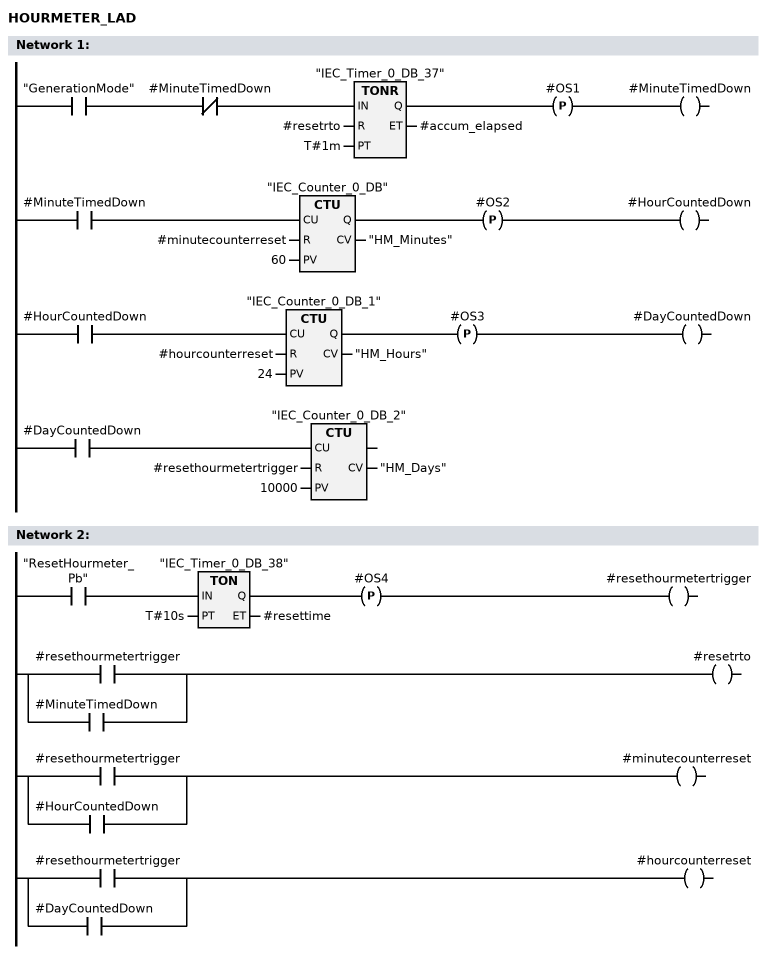
   "IEC_Timer_0_DB_37".TONR(IN := "GenerationMode" AND NOT #MinuteTimedDown,
                           R := #resetrto,
                           PT := T#1m,
                           ET => #accum_elapsed);
   #_w1 := "IEC_Timer_0_DB_37".Q AND NOT #OS1;   // rising edge
   #OS1 := "IEC_Timer_0_DB_37".Q;
   #MinuteTimedDown := #_w1;
   "IEC_Counter_0_DB".CTU(CU := #MinuteTimedDown, R := #minutecounterreset, PV := 60, CV => "HM_Minutes");
   #_w2 := "IEC_Counter_0_DB".Q AND NOT #OS2;   // rising edge
   #OS2 := "IEC_Counter_0_DB".Q;
   #HourCountedDown := #_w2;
   "IEC_Counter_0_DB_1".CTU(CU := #HourCountedDown, R := #hourcounterreset, PV := 24, CV => "HM_Hours");
   #_w3 := "IEC_Counter_0_DB_1".Q AND NOT #OS3;   // rising edge
   #OS3 := "IEC_Counter_0_DB_1".Q;
   #DayCountedDown := #_w3;
   "IEC_Counter_0_DB_2".CTU(CU := #DayCountedDown, R := #resethourmetertrigger, PV := 10000, CV => "HM_Days");
END_REGION

REGION Network 2
   "IEC_Timer_0_DB_38".TON(IN := "ResetHourmeter_Pb", PT := T#10s, ET => #resettime);
   #_w1 := "IEC_Timer_0_DB_38".Q AND NOT #OS4;   // rising edge
   #OS4 := "IEC_Timer_0_DB_38".Q;
   #resethourmetertrigger := #_w1;
   #resetrto := #resethourmetertrigger OR #MinuteTimedDown;
   #minutecounterreset := #resethourmetertrigger OR #HourCountedDown;
   #hourcounterreset := #resethourmetertrigger OR #DayCountedDown;
END_REGION
END_FUNCTION_BLOCK

FUNCTION_BLOCK "HOURMETER_FBD"   // FB20, FBD
{ S7_Optimized_Access := 'TRUE' }
VERSION : 0.1
   VAR
      OS1 : Bool;
      OS2 : Bool;
      OS3 : Bool;
      OS4 : Bool;
      rtotimerreset : Bool;
      minutecounterreset : Bool;
      hourcounterreset : Bool;
      hourmeterresettrigger : Bool;
      accumulatedtime : Time;
      minutetimeddown : Bool;
      hourcounteddown : Bool;
      daycounteddown : Bool;
   END_VAR
   VAR_TEMP   // added for the SCL form of the ladder/FBD networks
      _w1 : Bool;
      _w2 : Bool;
      _w3 : Bool;
   END_VAR
BEGIN

REGION Network 1
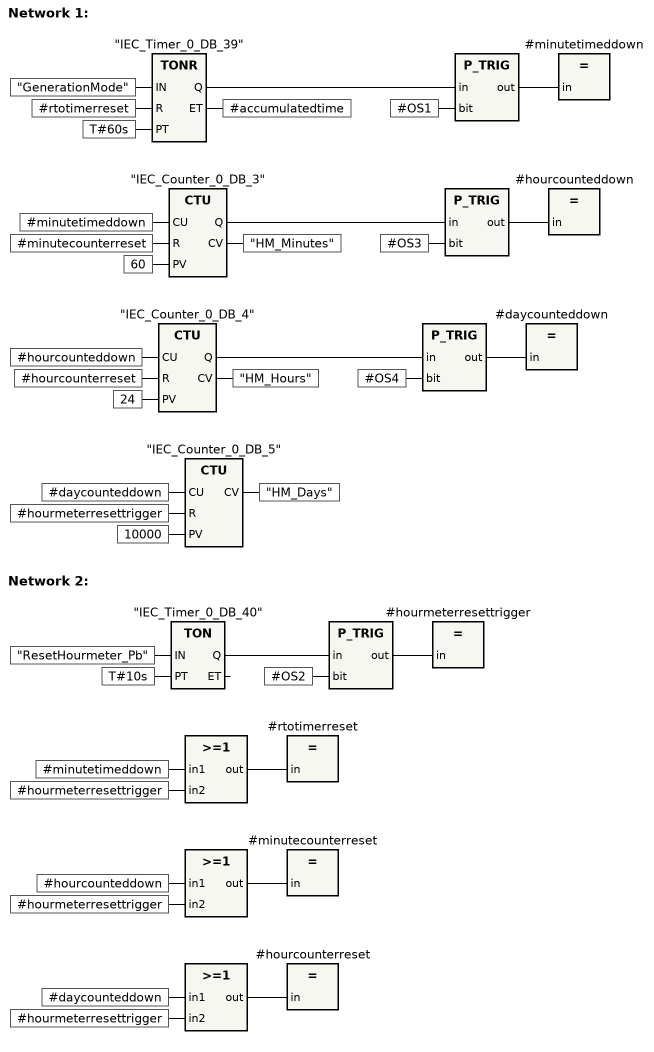
   "IEC_Timer_0_DB_39".TONR(IN := "GenerationMode", R := #rtotimerreset, PT := T#60s, ET => #accumulatedtime);
   #_w1 := "IEC_Timer_0_DB_39".Q AND NOT #OS1;   // rising edge
   #OS1 := "IEC_Timer_0_DB_39".Q;
   #minutetimeddown := #_w1;
   "IEC_Counter_0_DB_3".CTU(CU := #minutetimeddown, R := #minutecounterreset, PV := 60, CV => "HM_Minutes");
   #_w2 := "IEC_Counter_0_DB_3".Q AND NOT #OS3;   // rising edge
   #OS3 := "IEC_Counter_0_DB_3".Q;
   #hourcounteddown := #_w2;
   "IEC_Counter_0_DB_4".CTU(CU := #hourcounteddown, R := #hourcounterreset, PV := 24, CV => "HM_Hours");
   #_w3 := "IEC_Counter_0_DB_4".Q AND NOT #OS4;   // rising edge
   #OS4 := "IEC_Counter_0_DB_4".Q;
   #daycounteddown := #_w3;
   "IEC_Counter_0_DB_5".CTU(CU := #daycounteddown, R := #hourmeterresettrigger, PV := 10000, CV => "HM_Days");
END_REGION

REGION Network 2
   "IEC_Timer_0_DB_40".TON(IN := "ResetHourmeter_Pb", PT := T#10s);
   #_w1 := "IEC_Timer_0_DB_40".Q AND NOT #OS2;   // rising edge
   #OS2 := "IEC_Timer_0_DB_40".Q;
   #hourmeterresettrigger := #_w1;
   #rtotimerreset := #minutetimeddown OR #hourmeterresettrigger;
   #minutecounterreset := #hourcounteddown OR #hourmeterresettrigger;
   #hourcounterreset := #daycounteddown OR #hourmeterresettrigger;
END_REGION
END_FUNCTION_BLOCK

FUNCTION_BLOCK "HOURMETER_SCL"   // FB21, SCL
{ S7_Optimized_Access := 'TRUE' }
VERSION : 0.1
   VAR
      rtotimerreset : Bool;
      minutecounterreset : Bool;
      hourcounterreset : Bool;
      hourmeterresettrigger : Bool;
      accumulatedtime : Time;
      minutetimeddown : Bool;
      hourcounteddown : Bool;
      daycounteddown : Bool;
   END_VAR
BEGIN
   IF "GenerationMode" THEN
       "IEC_Timer_0_DB_41".TONR(IN := TRUE,
                                R := #rtotimerreset,
                                PT := T#60s,
                                Q => #minutetimeddown,
                                ET => #accumulatedtime);
   END_IF;

   IF #minutetimeddown THEN
       RESET_TIMER("IEC_Timer_0_DB_41");
   END_IF;

   "IEC_Counter_0_DB_6".CTU(CU:=#minutetimeddown,
                            R:=#minutecounterreset,
                            PV:=60,
                            Q=>#hourcounteddown,
                            CV=>"HM_Minutes");

   "IEC_Counter_0_DB_7".CTU(CU:=#hourcounteddown,
                            R:=#hourcounterreset,
                            PV:=24,
                            Q=>#daycounteddown,
                            CV=>"HM_Hours");

   "IEC_Counter_0_DB_9".CTU(CU:=#daycounteddown,
                            R:=#hourmeterresettrigger,
                            PV:=10000,
                            CV=>"HM_Days");

   IF "ResetHourmeter_Pb" THEN
       "IEC_Timer_0_DB_42".TON(IN:=TRUE,
                               PT:=T#10s,
                               Q=>#hourmeterresettrigger);
   ELSE
       RESET_TIMER("IEC_Timer_0_DB_42");
   END_IF;

   IF #hourmeterresettrigger OR #minutetimeddown THEN
       #rtotimerreset := 1;
   ELSE
       #rtotimerreset := 0;
   END_IF;

   IF #hourmeterresettrigger OR #hourcounteddown THEN
       #minutecounterreset := 1;
   ELSE
       #minutecounterreset := 0;
   END_IF;

   IF #hourmeterresettrigger OR #daycounteddown THEN
       #hourcounterreset := 1;
   ELSE
       #hourcounterreset := 0;
   END_IF;
END_FUNCTION_BLOCK

FUNCTION_BLOCK "HOURMETER_STL"   // FB22, STL
{ S7_Optimized_Access := 'TRUE' }
VERSION : 0.1
   VAR
      hourmeterresettrigger : Bool;
      minutecounterreset : Bool;
      hourcounterreset : Bool;
      minutetimeddown : Bool;
      hourcounteddown : Bool;
      daycounteddown : Bool;
      accumulatedtime : Time;
      rtotimerreset : Bool;
   END_VAR
   VAR_TEMP
      toomanydays : Bool;
      acctime : Time;
   END_VAR
BEGIN

REGION Network 1
         A     "GenerationMode";
         JC    RTOtimer;
         CLR;
         JU    EndOfLine;

   RTOtimer:CALL  TONR, "IEC_Timer_0_DB_43"
         ( IN := TRUE,
           R  := #rtotimerreset,
           PT := T#1m,
           Q  := #minutetimeddown,
           ET := #accumulatedtime
         );

         CALL  CTU, "IEC_Counter_0_DB_10"
         ( CU := #minutetimeddown,
           R  := #minutecounterreset,
           PV := 60,
           Q  := #hourcounteddown,
           CV := "HM_Minutes"
         );

         CALL  CTU, "IEC_Counter_0_DB_11"
         ( CU := #hourcounteddown,
           R  := #hourcounterreset,
           PV := 24,
           Q  := #daycounteddown,
           CV := "HM_Hours"
         );

         CALL  CTU, "IEC_Counter_0_DB_12"
         ( CU := #daycounteddown,
           R  := #hourmeterresettrigger,
           PV := 10000,
           Q  := #toomanydays,
           CV := "HM_Days"
         );

         JU    ResetEvaluate;

   ResetEvaluate:CLR;
         A     "ResetHourmeter_Pb";
         JC    ResetHourmeter;
         CALL  RESET_TIMER
         ( "TIMER" := "IEC_Timer_0_DB_44"
         );
         JU    EndOfLine;

   ResetHourmeter:CALL  TON, "IEC_Timer_0_DB_44"
         ( IN := TRUE,
           PT := T#10s,
           Q  := #hourmeterresettrigger,
           ET := #acctime
         );


   EndOfLine:A     #hourmeterresettrigger;
         O     #minutetimeddown;
         =     #rtotimerreset;
         CLR;
         A     #hourmeterresettrigger;
         O     #hourcounteddown;
         =     #minutecounterreset;
         CLR;
         A     #hourmeterresettrigger;
         O     #daycounteddown;
         =     #hourcounterreset;
         CLR;
         NOT;
         R     #hourmeterresettrigger;
END_REGION
END_FUNCTION_BLOCK

FUNCTION "SCP" : Void   // FC1, FBD
{ S7_Optimized_Access := 'TRUE' }
VERSION : 0.1
   VAR_INPUT
      Input_Min : Int;
      Input_Signal : Int;
      Input_Max : Int;
      Output_Min : Int;
      Output_Max : Int;
   END_VAR
   VAR_OUTPUT
      SV : Int;
   END_VAR
   VAR_TEMP
      tv : Real;
   END_VAR
BEGIN

REGION Network 1
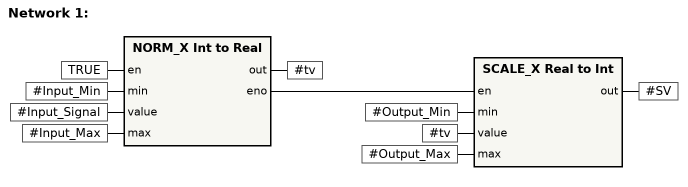
   IF TRUE THEN
       #tv := NORM_X(MIN := #Input_Min, VALUE := #Input_Signal, MAX := #Input_Max);
       #SV := SCALE_X(MIN := #Output_Min, VALUE := #tv, MAX := #Output_Max);
   END_IF;
END_REGION
END_FUNCTION

FUNCTION "CONVERTTIME" : Void   // FC2, FBD
{ S7_Optimized_Access := 'TRUE' }
VERSION : 0.1
   VAR_INPUT
      Int1 : Int;
   END_VAR
   VAR_OUTPUT
      Time1 : Time;
   END_VAR
   VAR_TEMP
      tv : Int;
   END_VAR
BEGIN

REGION Network 1
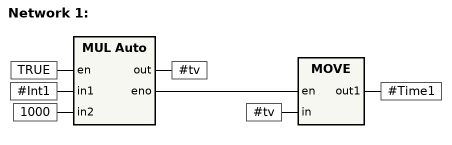
   IF TRUE THEN
       #tv := #Int1 * 1000;
       #Time1 := #tv;
   END_IF;
END_REGION
END_FUNCTION

ORGANIZATION_BLOCK "Main"   // OB1, LAD, ProgramCycle
TITLE = "Main Program Sweep (Cycle)"
{ S7_Optimized_Access := 'TRUE' }
VERSION : 0.1
   VAR_INPUT
      Initial_Call : Bool;   // Initial call of this OB
      Remanence : Bool;   // =True, if remanent data are available
   END_VAR
   VAR_TEMP
      SequenceInit : Bool;
      InitSequence : Bool;
   END_VAR
   VAR_TEMP   // added for the SCL form of the ladder/FBD networks
      _w1 : Bool;
      _w2 : Bool;
      _w3 : Bool;
      _w4 : Bool;
   END_VAR
BEGIN

REGION Network 1
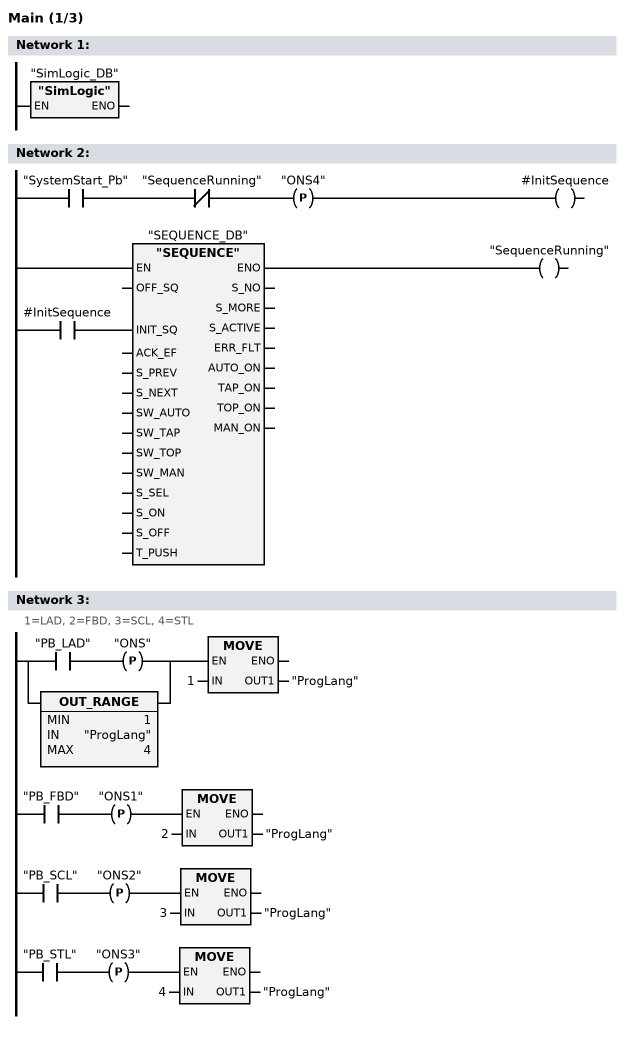
   RUNG wire#powerrail
      "SimLogic_DB"()
   END_RUNG
   // the same network as SCL:
   "SimLogic_DB"();   // "SimLogic"
END_REGION

REGION Network 2
   RUNG wire#powerrail
      Contact( "SystemStart_Pb" )
      I_Contact( "SequenceRunning" )
      P_Trig( "ONS4" )
      Coil( #InitSequence )
   END_RUNG
   RUNG wire#powerrail
      "SEQUENCE_DB"(INIT_SQ := wire#w1, OFF_SQ :=, ACK_EF :=, S_PREV :=, S_NEXT :=, SW_AUTO :=, SW_TAP :=, SW_TOP :=, SW_MAN :=, S_SEL :=, S_ON :=, S_OFF :=, T_PUSH :=, S_NO =>, S_MORE =>, S_ACTIVE =>, ERR_FLT =>, AUTO_ON =>, TAP_ON =>, TOP_ON =>, MAN_ON =>)
      Coil( "SequenceRunning" )
   END_RUNG
   RUNG wire#powerrail
      Contact( #InitSequence )
   END_RUNG wire#w1
   // the same network as SCL:
   #_w1 := "SystemStart_Pb" AND NOT "SequenceRunning";
   #_w2 := #_w1 AND NOT "ONS4";   // rising edge
   "ONS4" := #_w1;
   #InitSequence := #_w2;
   "SEQUENCE_DB"(INIT_SQ := #InitSequence, ENO => #_w3);   // "SEQUENCE"
   "SequenceRunning" := #_w3;
END_REGION

REGION Network 3
   // 1=LAD, 2=FBD, 3=SCL, 4=STL
   #_w1 := "PB_LAD" AND NOT "ONS";   // rising edge
   "ONS" := "PB_LAD";
   IF #_w1 OR ("ProgLang" < 1) OR ("ProgLang" > 4) THEN "ProgLang" := 1; END_IF;
   #_w2 := "PB_FBD" AND NOT "ONS1";   // rising edge
   "ONS1" := "PB_FBD";
   IF #_w2 THEN "ProgLang" := 2; END_IF;
   #_w3 := "PB_SCL" AND NOT "ONS2";   // rising edge
   "ONS2" := "PB_SCL";
   IF #_w3 THEN "ProgLang" := 3; END_IF;
   #_w4 := "PB_STL" AND NOT "ONS3";   // rising edge
   "ONS3" := "PB_STL";
   IF #_w4 THEN "ProgLang" := 4; END_IF;
END_REGION

REGION Network 4
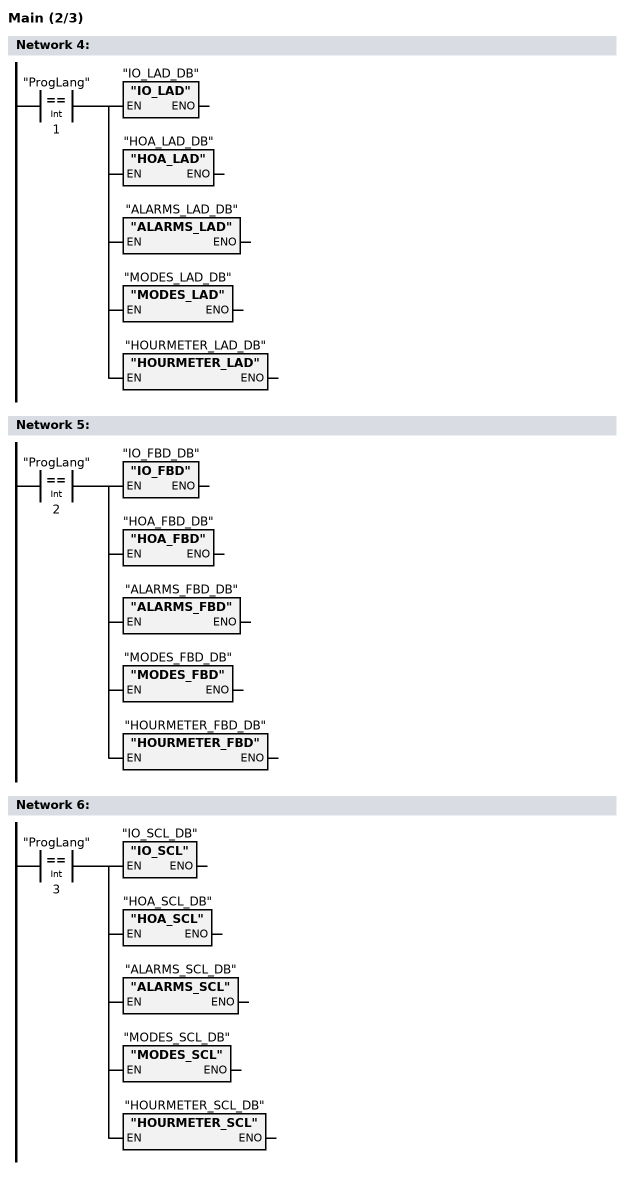
   RUNG wire#powerrail
      { S7_Templates := "SrcType := Int" } EQ_Contact(in1 := "ProgLang", in2 := 1)
      wire#w1
      "IO_LAD_DB"()
   END_RUNG
   RUNG wire#w1
      "HOA_LAD_DB"()
   END_RUNG
   RUNG wire#w1
      "ALARMS_LAD_DB"()
   END_RUNG
   RUNG wire#w1
      "MODES_LAD_DB"()
   END_RUNG
   RUNG wire#w1
      "HOURMETER_LAD_DB"()
   END_RUNG
   // the same network as SCL:
   #_w1 := "ProgLang" = 1;
   IF #_w1 THEN
       "IO_LAD_DB"();   // "IO_LAD"
       "HOA_LAD_DB"();   // "HOA_LAD"
       "ALARMS_LAD_DB"();   // "ALARMS_LAD"
       "MODES_LAD_DB"();   // "MODES_LAD"
       "HOURMETER_LAD_DB"();   // "HOURMETER_LAD"
   END_IF;
END_REGION

REGION Network 5
   RUNG wire#powerrail
      { S7_Templates := "SrcType := Int" } EQ_Contact(in1 := "ProgLang", in2 := 2)
      wire#w1
      "IO_FBD_DB"()
   END_RUNG
   RUNG wire#w1
      "HOA_FBD_DB"()
   END_RUNG
   RUNG wire#w1
      "ALARMS_FBD_DB"()
   END_RUNG
   RUNG wire#w1
      "MODES_FBD_DB"()
   END_RUNG
   RUNG wire#w1
      "HOURMETER_FBD_DB"()
   END_RUNG
   // the same network as SCL:
   #_w1 := "ProgLang" = 2;
   IF #_w1 THEN
       "IO_FBD_DB"();   // "IO_FBD"
       "HOA_FBD_DB"();   // "HOA_FBD"
       "ALARMS_FBD_DB"();   // "ALARMS_FBD"
       "MODES_FBD_DB"();   // "MODES_FBD"
       "HOURMETER_FBD_DB"();   // "HOURMETER_FBD"
   END_IF;
END_REGION

REGION Network 6
   RUNG wire#powerrail
      { S7_Templates := "SrcType := Int" } EQ_Contact(in1 := "ProgLang", in2 := 3)
      wire#w1
      "IO_SCL_DB"()
   END_RUNG
   RUNG wire#w1
      "HOA_SCL_DB"()
   END_RUNG
   RUNG wire#w1
      "ALARMS_SCL_DB"()
   END_RUNG
   RUNG wire#w1
      "MODES_SCL_DB"()
   END_RUNG
   RUNG wire#w1
      "HOURMETER_SCL_DB"()
   END_RUNG
   // the same network as SCL:
   #_w1 := "ProgLang" = 3;
   IF #_w1 THEN
       "IO_SCL_DB"();   // "IO_SCL"
       "HOA_SCL_DB"();   // "HOA_SCL"
       "ALARMS_SCL_DB"();   // "ALARMS_SCL"
       "MODES_SCL_DB"();   // "MODES_SCL"
       "HOURMETER_SCL_DB"();   // "HOURMETER_SCL"
   END_IF;
END_REGION

REGION Network 7
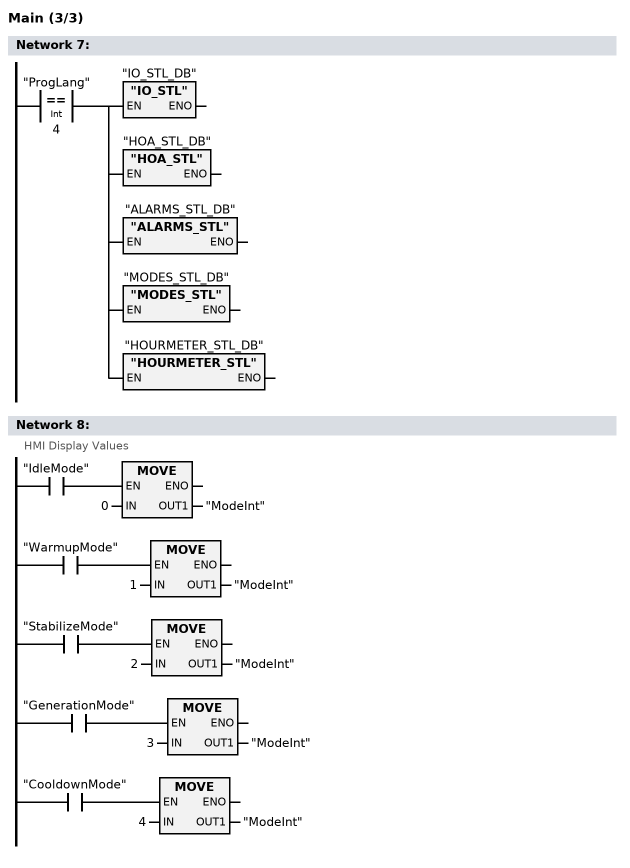
   RUNG wire#powerrail
      { S7_Templates := "SrcType := Int" } EQ_Contact(in1 := "ProgLang", in2 := 4)
      wire#w1
      "IO_STL_DB"()
   END_RUNG
   RUNG wire#w1
      "HOA_STL_DB"()
   END_RUNG
   RUNG wire#w1
      "ALARMS_STL_DB"()
   END_RUNG
   RUNG wire#w1
      "MODES_STL_DB"()
   END_RUNG
   RUNG wire#w1
      "HOURMETER_STL_DB"()
   END_RUNG
   // the same network as SCL:
   #_w1 := "ProgLang" = 4;
   IF #_w1 THEN
       "IO_STL_DB"();   // "IO_STL"
       "HOA_STL_DB"();   // "HOA_STL"
       "ALARMS_STL_DB"();   // "ALARMS_STL"
       "MODES_STL_DB"();   // "MODES_STL"
       "HOURMETER_STL_DB"();   // "HOURMETER_STL"
   END_IF;
END_REGION

REGION Network 8
   // HMI Display Values
   RUNG wire#powerrail
      Contact( "IdleMode" )
      Move(in := 0, out1 => "ModeInt")
   END_RUNG
   RUNG wire#powerrail
      Contact( "WarmupMode" )
      Move(in := 1, out1 => "ModeInt")
   END_RUNG
   RUNG wire#powerrail
      Contact( "StabilizeMode" )
      Move(in := 2, out1 => "ModeInt")
   END_RUNG
   RUNG wire#powerrail
      Contact( "GenerationMode" )
      Move(in := 3, out1 => "ModeInt")
   END_RUNG
   RUNG wire#powerrail
      Contact( "CooldownMode" )
      Move(in := 4, out1 => "ModeInt")
   END_RUNG
   // the same network as SCL:
   IF "IdleMode" THEN "ModeInt" := 0; END_IF;
   IF "WarmupMode" THEN "ModeInt" := 1; END_IF;
   IF "StabilizeMode" THEN "ModeInt" := 2; END_IF;
   IF "GenerationMode" THEN "ModeInt" := 3; END_IF;
   IF "CooldownMode" THEN "ModeInt" := 4; END_IF;
END_REGION
END_ORGANIZATION_BLOCK

ORGANIZATION_BLOCK "PID"   // OB31, LAD, CyclicInterrupt
{ S7_Optimized_Access := 'TRUE' }
VERSION : 0.1
   VAR_INPUT
      Initial_Call : Bool;   // Initial call of this OB
      Event_Count : Int;   // Events discarded
   END_VAR
   VAR_TEMP
      Bsp : Real;
      Vsp : Real;
      BaffleHandTrigger : Bool;
      BaffleOffTrigger : Bool;
      VFDHandTrigger : Bool;
      VFDOffTrigger : Bool;
      BaffleAutoTrigger : Bool;
      VFDautoTrigger : Bool;
   END_VAR
   VAR_TEMP   // added for the SCL form of the ladder/FBD networks
      _w1 : Bool;
      _w2 : Bool;
      _w3 : Bool;
      _w4 : Bool;
      _w5 : Bool;
      _w6 : Bool;
      _w7 : Bool;
   END_VAR
BEGIN

REGION Network 1
   // High Oil Flow Alarm Handling
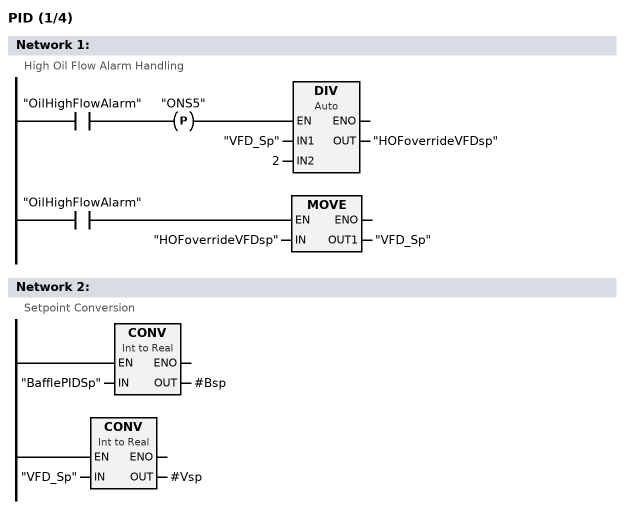
   RUNG wire#powerrail
      Contact( "OilHighFlowAlarm" )
      P_Trig( "ONS5" )
      Div(in1 := "VFD_Sp", in2 := 2, out => "HOFoverrideVFDsp")
   END_RUNG
   RUNG wire#powerrail
      Contact( "OilHighFlowAlarm" )
      Move(in := "HOFoverrideVFDsp", out1 => "VFD_Sp")
   END_RUNG
   // the same network as SCL:
   #_w1 := "OilHighFlowAlarm" AND NOT "ONS5";   // rising edge
   "ONS5" := "OilHighFlowAlarm";
   IF #_w1 THEN "HOFoverrideVFDsp" := "VFD_Sp" / 2; END_IF;
   IF "OilHighFlowAlarm" THEN "VFD_Sp" := "HOFoverrideVFDsp"; END_IF;
END_REGION

REGION Network 2
   // Setpoint Conversion
   RUNG wire#powerrail
      { S7_Templates := "[SrcType := Int, DestType := Real]" } Convert(in := "BafflePIDSp", out => #Bsp)
   END_RUNG
   RUNG wire#powerrail
      { S7_Templates := "[SrcType := Int, DestType := Real]" } Convert(in := "VFD_Sp", out => #Vsp)
   END_RUNG
   // the same network as SCL:
   #Bsp := INT_TO_REAL("BafflePIDSp");
   #Vsp := INT_TO_REAL("VFD_Sp");
END_REGION

REGION Network 3
   // Baffle HOA
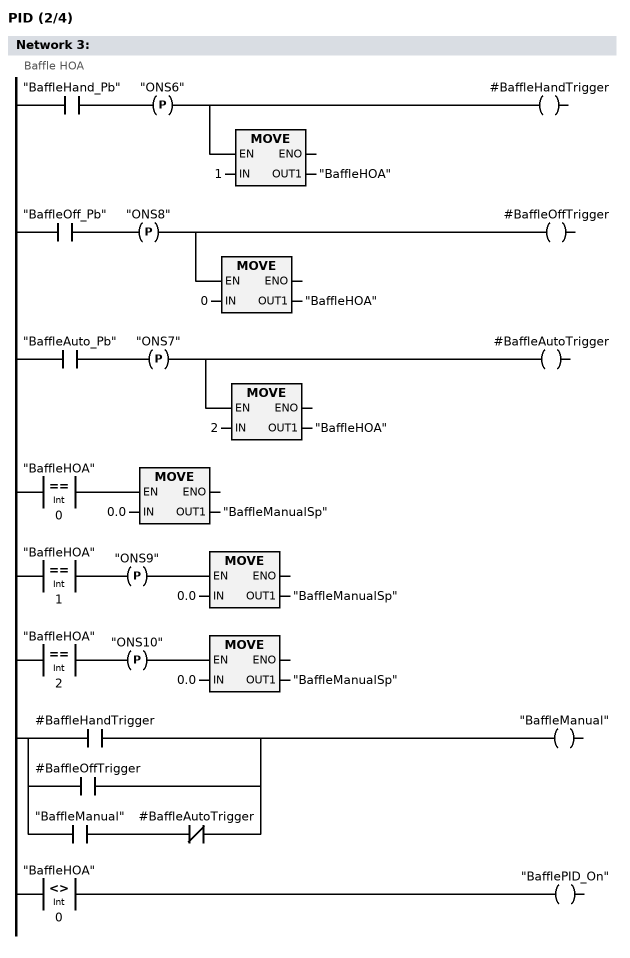
   RUNG wire#powerrail
      Contact( "BaffleHand_Pb" )
      P_Trig( "ONS6" )
      wire#w1
      Coil( #BaffleHandTrigger )
   END_RUNG
   RUNG wire#w1
      Move(in := 1, out1 => "BaffleHOA")
   END_RUNG
   RUNG wire#powerrail
      Contact( "BaffleOff_Pb" )
      P_Trig( "ONS8" )
      wire#w2
      Coil( #BaffleOffTrigger )
   END_RUNG
   RUNG wire#w2
      Move(in := 0, out1 => "BaffleHOA")
   END_RUNG
   RUNG wire#powerrail
      Contact( "BaffleAuto_Pb" )
      P_Trig( "ONS7" )
      wire#w3
      Coil( #BaffleAutoTrigger )
   END_RUNG
   RUNG wire#w3
      Move(in := 2, out1 => "BaffleHOA")
   END_RUNG
   RUNG wire#powerrail
      { S7_Templates := "SrcType := Int" } EQ_Contact(in1 := "BaffleHOA", in2 := 0)
      Move(in := 0.0, out1 => "BaffleManualSp")
   END_RUNG
   RUNG wire#powerrail
      { S7_Templates := "SrcType := Int" } EQ_Contact(in1 := "BaffleHOA", in2 := 1)
      P_Trig( "ONS9" )
      Move(in := 0.0, out1 => "BaffleManualSp")
   END_RUNG
   RUNG wire#powerrail
      { S7_Templates := "SrcType := Int" } EQ_Contact(in1 := "BaffleHOA", in2 := 2)
      P_Trig( "ONS10" )
      Move(in := 0.0, out1 => "BaffleManualSp")
   END_RUNG
   RUNG wire#powerrail
      Contact( #BaffleHandTrigger )
      wire#w4
      Coil( "BaffleManual" )
   END_RUNG
   RUNG wire#powerrail
      Contact( #BaffleOffTrigger )
   END_RUNG wire#w4
   RUNG wire#powerrail
      Contact( "BaffleManual" )
      I_Contact( #BaffleAutoTrigger )
   END_RUNG wire#w4
   RUNG wire#powerrail
      { S7_Templates := "SrcType := Int" } NE_Contact(in1 := "BaffleHOA", in2 := 0)
      Coil( "BafflePID_On" )
   END_RUNG
   // the same network as SCL:
   #_w1 := "BaffleHand_Pb" AND NOT "ONS6";   // rising edge
   "ONS6" := "BaffleHand_Pb";
   #BaffleHandTrigger := #_w1;
   IF #_w1 THEN "BaffleHOA" := 1; END_IF;
   #_w2 := "BaffleOff_Pb" AND NOT "ONS8";   // rising edge
   "ONS8" := "BaffleOff_Pb";
   #BaffleOffTrigger := #_w2;
   IF #_w2 THEN "BaffleHOA" := 0; END_IF;
   #_w3 := "BaffleAuto_Pb" AND NOT "ONS7";   // rising edge
   "ONS7" := "BaffleAuto_Pb";
   #BaffleAutoTrigger := #_w3;
   IF #_w3 THEN "BaffleHOA" := 2; END_IF;
   IF "BaffleHOA" = 0 THEN "BaffleManualSp" := 0.0; END_IF;
   #_w4 := "BaffleHOA" = 1;
   #_w5 := #_w4 AND NOT "ONS9";   // rising edge
   "ONS9" := #_w4;
   IF #_w5 THEN "BaffleManualSp" := 0.0; END_IF;
   #_w6 := "BaffleHOA" = 2;
   #_w7 := #_w6 AND NOT "ONS10";   // rising edge
   "ONS10" := #_w6;
   IF #_w7 THEN "BaffleManualSp" := 0.0; END_IF;
   "BaffleManual" := #BaffleHandTrigger OR #BaffleOffTrigger OR ("BaffleManual" AND NOT #BaffleAutoTrigger);
   "BafflePID_On" := "BaffleHOA" <> 0;
END_REGION

REGION Network 4
   // VFD HOA